(* Logix 5000 project; controller OWF Emulate 5570 rev 30.12; software revision 30.00; part 8 of 21 *)
(* tags used below, declared in another part *)
   OWF_Add_c : DINT;
   OWF_Input : DINT[16];
   OWF_Result : DINT[17];
(* MainProgram, continued *)

   	End_If;
   	If OWF_Input[7].[22] Then
   		OWF_Result[0]:=OWF_Result[0] + 480646434+OWF_Add_c;
   		OWF_Add_c.0:=OWF_Result[0].31;
   		OWF_Result[0].31:=0;
   		OWF_Result[1]:=OWF_Result[1] + 114796889+OWF_Add_c;
   		OWF_Add_c.1:=OWF_Result[1].31;
   		OWF_Result[1].31:=0;
   		OWF_Result[2]:=OWF_Result[2] + 808245238+OWF_Add_c;
   		OWF_Add_c.2:=OWF_Result[2].31;
   		OWF_Result[2].31:=0;
   		OWF_Result[3]:=OWF_Result[3] + 1045553390+OWF_Add_c;
   		OWF_Add_c.3:=OWF_Result[3].31;
   		OWF_Result[3].31:=0;
   		OWF_Result[4]:=OWF_Result[4] + 1347272097+OWF_Add_c;
   		OWF_Add_c.4:=OWF_Result[4].31;
   		OWF_Result[4].31:=0;
   		OWF_Result[5]:=OWF_Result[5] + 212393883+OWF_Add_c;
   		OWF_Add_c.5:=OWF_Result[5].31;
   		OWF_Result[5].31:=0;
   		OWF_Result[6]:=OWF_Result[6] + 833811458+OWF_Add_c;
   		OWF_Add_c.6:=OWF_Result[6].31;
   		OWF_Result[6].31:=0;
   		OWF_Result[7]:=OWF_Result[7] + 657498953+OWF_Add_c;
   		OWF_Add_c.7:=OWF_Result[7].31;
   		OWF_Result[7].31:=0;
   		OWF_Result[8]:=OWF_Result[8] + 1633172185+OWF_Add_c;
   		OWF_Add_c.8:=OWF_Result[8].31;
   		OWF_Result[8].31:=0;
   		OWF_Result[9]:=OWF_Result[9] + 109189510+OWF_Add_c;
   		OWF_Add_c.9:=OWF_Result[9].31;
   		OWF_Result[9].31:=0;
   		OWF_Result[10]:=OWF_Result[10] + 1987125799+OWF_Add_c;
   		OWF_Add_c.10:=OWF_Result[10].31;
   		OWF_Result[10].31:=0;
   		OWF_Result[11]:=OWF_Result[11] + 790477840+OWF_Add_c;
   		OWF_Add_c.11:=OWF_Result[11].31;
   		OWF_Result[11].31:=0;
   		OWF_Result[12]:=OWF_Result[12] + 1317536711+OWF_Add_c;
   		OWF_Add_c.12:=OWF_Result[12].31;
   		OWF_Result[12].31:=0;
   	End_If;
   	If OWF_Input[7].[23] Then
   		OWF_Result[0]:=OWF_Result[0] + 740299143+OWF_Add_c;
   		OWF_Add_c.0:=OWF_Result[0].31;
   		OWF_Result[0].31:=0;
   		OWF_Result[1]:=OWF_Result[1] + 289363045+OWF_Add_c;
   		OWF_Add_c.1:=OWF_Result[1].31;
   		OWF_Result[1].31:=0;
   		OWF_Result[2]:=OWF_Result[2] + 506118578+OWF_Add_c;
   		OWF_Add_c.2:=OWF_Result[2].31;
   		OWF_Result[2].31:=0;
   		OWF_Result[3]:=OWF_Result[3] + 1440714184+OWF_Add_c;
   		OWF_Add_c.3:=OWF_Result[3].31;
   		OWF_Result[3].31:=0;
   		OWF_Result[4]:=OWF_Result[4] + 1773567421+OWF_Add_c;
   		OWF_Add_c.4:=OWF_Result[4].31;
   		OWF_Result[4].31:=0;
   		OWF_Result[5]:=OWF_Result[5] + 1795348463+OWF_Add_c;
   		OWF_Add_c.5:=OWF_Result[5].31;
   		OWF_Result[5].31:=0;
   		OWF_Result[6]:=OWF_Result[6] + 1980498485+OWF_Add_c;
   		OWF_Add_c.6:=OWF_Result[6].31;
   		OWF_Result[6].31:=0;
   		OWF_Result[7]:=OWF_Result[7] + 308789052+OWF_Add_c;
   		OWF_Add_c.7:=OWF_Result[7].31;
   		OWF_Result[7].31:=0;
   		OWF_Result[8]:=OWF_Result[8] + 1048758798+OWF_Add_c;
   		OWF_Add_c.8:=OWF_Result[8].31;
   		OWF_Result[8].31:=0;
   		OWF_Result[9]:=OWF_Result[9] + 916377049+OWF_Add_c;
   		OWF_Add_c.9:=OWF_Result[9].31;
   		OWF_Result[9].31:=0;
   		OWF_Result[10]:=OWF_Result[10] + 502789876+OWF_Add_c;
   		OWF_Add_c.10:=OWF_Result[10].31;
   		OWF_Result[10].31:=0;
   		OWF_Result[11]:=OWF_Result[11] + 629743481+OWF_Add_c;
   		OWF_Add_c.11:=OWF_Result[11].31;
   		OWF_Result[11].31:=0;
   		OWF_Result[12]:=OWF_Result[12] + 1676079784+OWF_Add_c;
   		OWF_Add_c.12:=OWF_Result[12].31;
   		OWF_Result[12].31:=0;
   	End_If;
   	If OWF_Input[7].[24] Then
   		OWF_Result[0]:=OWF_Result[0] + 978983842+OWF_Add_c;
   		OWF_Add_c.0:=OWF_Result[0].31;
   		OWF_Result[0].31:=0;
   		OWF_Result[1]:=OWF_Result[1] + 184076912+OWF_Add_c;
   		OWF_Add_c.1:=OWF_Result[1].31;
   		OWF_Result[1].31:=0;
   		OWF_Result[2]:=OWF_Result[2] + 18075719+OWF_Add_c;
   		OWF_Add_c.2:=OWF_Result[2].31;
   		OWF_Result[2].31:=0;
   		OWF_Result[3]:=OWF_Result[3] + 1672505732+OWF_Add_c;
   		OWF_Add_c.3:=OWF_Result[3].31;
   		OWF_Result[3].31:=0;
   		OWF_Result[4]:=OWF_Result[4] + 1803238491+OWF_Add_c;
   		OWF_Add_c.4:=OWF_Result[4].31;
   		OWF_Result[4].31:=0;
   		OWF_Result[5]:=OWF_Result[5] + 1332716281+OWF_Add_c;
   		OWF_Add_c.5:=OWF_Result[5].31;
   		OWF_Result[5].31:=0;
   		OWF_Result[6]:=OWF_Result[6] + 633027607+OWF_Add_c;
   		OWF_Add_c.6:=OWF_Result[6].31;
   		OWF_Result[6].31:=0;
   		OWF_Result[7]:=OWF_Result[7] + 1542211604+OWF_Add_c;
   		OWF_Add_c.7:=OWF_Result[7].31;
   		OWF_Result[7].31:=0;
   		OWF_Result[8]:=OWF_Result[8] + 716891059+OWF_Add_c;
   		OWF_Add_c.8:=OWF_Result[8].31;
   		OWF_Result[8].31:=0;
   		OWF_Result[9]:=OWF_Result[9] + 1337341351+OWF_Add_c;
   		OWF_Add_c.9:=OWF_Result[9].31;
   		OWF_Result[9].31:=0;
   		OWF_Result[10]:=OWF_Result[10] + 1718317461+OWF_Add_c;
   		OWF_Add_c.10:=OWF_Result[10].31;
   		OWF_Result[10].31:=0;
   		OWF_Result[11]:=OWF_Result[11] + 759267344+OWF_Add_c;
   		OWF_Add_c.11:=OWF_Result[11].31;
   		OWF_Result[11].31:=0;
   		OWF_Result[12]:=OWF_Result[12] + 1222721366+OWF_Add_c;
   		OWF_Add_c.12:=OWF_Result[12].31;
   		OWF_Result[12].31:=0;
   	End_If;
   	If OWF_Input[7].[25] Then
   		OWF_Result[0]:=OWF_Result[0] + 1210573640+OWF_Add_c;
   		OWF_Add_c.0:=OWF_Result[0].31;
   		OWF_Result[0].31:=0;
   		OWF_Result[1]:=OWF_Result[1] + 1066502865+OWF_Add_c;
   		OWF_Add_c.1:=OWF_Result[1].31;
   		OWF_Result[1].31:=0;
   		OWF_Result[2]:=OWF_Result[2] + 20470411+OWF_Add_c;
   		OWF_Add_c.2:=OWF_Result[2].31;
   		OWF_Result[2].31:=0;
   		OWF_Result[3]:=OWF_Result[3] + 526137192+OWF_Add_c;
   		OWF_Add_c.3:=OWF_Result[3].31;
   		OWF_Result[3].31:=0;
   		OWF_Result[4]:=OWF_Result[4] + 428761318+OWF_Add_c;
   		OWF_Add_c.4:=OWF_Result[4].31;
   		OWF_Result[4].31:=0;
   		OWF_Result[5]:=OWF_Result[5] + 666284081+OWF_Add_c;
   		OWF_Add_c.5:=OWF_Result[5].31;
   		OWF_Result[5].31:=0;
   		OWF_Result[6]:=OWF_Result[6] + 787646009+OWF_Add_c;
   		OWF_Add_c.6:=OWF_Result[6].31;
   		OWF_Result[6].31:=0;
   		OWF_Result[7]:=OWF_Result[7] + 1465565705+OWF_Add_c;
   		OWF_Add_c.7:=OWF_Result[7].31;
   		OWF_Result[7].31:=0;
   		OWF_Result[8]:=OWF_Result[8] + 2117689109+OWF_Add_c;
   		OWF_Add_c.8:=OWF_Result[8].31;
   		OWF_Result[8].31:=0;
   		OWF_Result[9]:=OWF_Result[9] + 1455398601+OWF_Add_c;
   		OWF_Add_c.9:=OWF_Result[9].31;
   		OWF_Result[9].31:=0;
   		OWF_Result[10]:=OWF_Result[10] + 732503870+OWF_Add_c;
   		OWF_Add_c.10:=OWF_Result[10].31;
   		OWF_Result[10].31:=0;
   		OWF_Result[11]:=OWF_Result[11] + 1389721484+OWF_Add_c;
   		OWF_Add_c.11:=OWF_Result[11].31;
   		OWF_Result[11].31:=0;
   		OWF_Result[12]:=OWF_Result[12] + 1051435137+OWF_Add_c;
   		OWF_Add_c.12:=OWF_Result[12].31;
   		OWF_Result[12].31:=0;
   	End_If;
   	If OWF_Input[7].[26] Then
   		OWF_Result[0]:=OWF_Result[0] + 1093740877+OWF_Add_c;
   		OWF_Add_c.0:=OWF_Result[0].31;
   		OWF_Result[0].31:=0;
   		OWF_Result[1]:=OWF_Result[1] + 1926933030+OWF_Add_c;
   		OWF_Add_c.1:=OWF_Result[1].31;
   		OWF_Result[1].31:=0;
   		OWF_Result[2]:=OWF_Result[2] + 2048297708+OWF_Add_c;
   		OWF_Add_c.2:=OWF_Result[2].31;
   		OWF_Result[2].31:=0;
   		OWF_Result[3]:=OWF_Result[3] + 1774994164+OWF_Add_c;
   		OWF_Add_c.3:=OWF_Result[3].31;
   		OWF_Result[3].31:=0;
   		OWF_Result[4]:=OWF_Result[4] + 100463613+OWF_Add_c;
   		OWF_Add_c.4:=OWF_Result[4].31;
   		OWF_Result[4].31:=0;
   		OWF_Result[5]:=OWF_Result[5] + 1811813667+OWF_Add_c;
   		OWF_Add_c.5:=OWF_Result[5].31;
   		OWF_Result[5].31:=0;
   		OWF_Result[6]:=OWF_Result[6] + 1209213066+OWF_Add_c;
   		OWF_Add_c.6:=OWF_Result[6].31;
   		OWF_Result[6].31:=0;
   		OWF_Result[7]:=OWF_Result[7] + 1269950558+OWF_Add_c;
   		OWF_Add_c.7:=OWF_Result[7].31;
   		OWF_Result[7].31:=0;
   		OWF_Result[8]:=OWF_Result[8] + 624695169+OWF_Add_c;
   		OWF_Add_c.8:=OWF_Result[8].31;
   		OWF_Result[8].31:=0;
   		OWF_Result[9]:=OWF_Result[9] + 1916749071+OWF_Add_c;
   		OWF_Add_c.9:=OWF_Result[9].31;
   		OWF_Result[9].31:=0;
   		OWF_Result[10]:=OWF_Result[10] + 1775084911+OWF_Add_c;
   		OWF_Add_c.10:=OWF_Result[10].31;
   		OWF_Result[10].31:=0;
   		OWF_Result[11]:=OWF_Result[11] + 1305211684+OWF_Add_c;
   		OWF_Add_c.11:=OWF_Result[11].31;
   		OWF_Result[11].31:=0;
   		OWF_Result[12]:=OWF_Result[12] + 546822773+OWF_Add_c;
   		OWF_Add_c.12:=OWF_Result[12].31;
   		OWF_Result[12].31:=0;
   	End_If;
   	If OWF_Input[7].[27] Then
   		OWF_Result[0]:=OWF_Result[0] + 859091503+OWF_Add_c;
   		OWF_Add_c.0:=OWF_Result[0].31;
   		OWF_Result[0].31:=0;
   		OWF_Result[1]:=OWF_Result[1] + 734881955+OWF_Add_c;
   		OWF_Add_c.1:=OWF_Result[1].31;
   		OWF_Result[1].31:=0;
   		OWF_Result[2]:=OWF_Result[2] + 2112245734+OWF_Add_c;
   		OWF_Add_c.2:=OWF_Result[2].31;
   		OWF_Result[2].31:=0;
   		OWF_Result[3]:=OWF_Result[3] + 821086543+OWF_Add_c;
   		OWF_Add_c.3:=OWF_Result[3].31;
   		OWF_Result[3].31:=0;
   		OWF_Result[4]:=OWF_Result[4] + 172634749+OWF_Add_c;
   		OWF_Add_c.4:=OWF_Result[4].31;
   		OWF_Result[4].31:=0;
   		OWF_Result[5]:=OWF_Result[5] + 1640326127+OWF_Add_c;
   		OWF_Add_c.5:=OWF_Result[5].31;
   		OWF_Result[5].31:=0;
   		OWF_Result[6]:=OWF_Result[6] + 90813347+OWF_Add_c;
   		OWF_Add_c.6:=OWF_Result[6].31;
   		OWF_Result[6].31:=0;
   		OWF_Result[7]:=OWF_Result[7] + 375324933+OWF_Add_c;
   		OWF_Add_c.7:=OWF_Result[7].31;
   		OWF_Result[7].31:=0;
   		OWF_Result[8]:=OWF_Result[8] + 734165162+OWF_Add_c;
   		OWF_Add_c.8:=OWF_Result[8].31;
   		OWF_Result[8].31:=0;
   		OWF_Result[9]:=OWF_Result[9] + 1211646497+OWF_Add_c;
   		OWF_Add_c.9:=OWF_Result[9].31;
   		OWF_Result[9].31:=0;
   		OWF_Result[10]:=OWF_Result[10] + 243057850+OWF_Add_c;
   		OWF_Add_c.10:=OWF_Result[10].31;
   		OWF_Result[10].31:=0;
   		OWF_Result[11]:=OWF_Result[11] + 2097424801+OWF_Add_c;
   		OWF_Add_c.11:=OWF_Result[11].31;
   		OWF_Result[11].31:=0;
   		OWF_Result[12]:=OWF_Result[12] + 609462236+OWF_Add_c;
   		OWF_Add_c.12:=OWF_Result[12].31;
   		OWF_Result[12].31:=0;
   	End_If;
   	If OWF_Input[7].[28] Then
   		OWF_Result[0]:=OWF_Result[0] + 1748630085+OWF_Add_c;
   		OWF_Add_c.0:=OWF_Result[0].31;
   		OWF_Result[0].31:=0;
   		OWF_Result[1]:=OWF_Result[1] + 218806354+OWF_Add_c;
   		OWF_Add_c.1:=OWF_Result[1].31;
   		OWF_Result[1].31:=0;
   		OWF_Result[2]:=OWF_Result[2] + 596066578+OWF_Add_c;
   		OWF_Add_c.2:=OWF_Result[2].31;
   		OWF_Result[2].31:=0;
   		OWF_Result[3]:=OWF_Result[3] + 1279944685+OWF_Add_c;
   		OWF_Add_c.3:=OWF_Result[3].31;
   		OWF_Result[3].31:=0;
   		OWF_Result[4]:=OWF_Result[4] + 798939716+OWF_Add_c;
   		OWF_Add_c.4:=OWF_Result[4].31;
   		OWF_Result[4].31:=0;
   		OWF_Result[5]:=OWF_Result[5] + 1193007422+OWF_Add_c;
   		OWF_Add_c.5:=OWF_Result[5].31;
   		OWF_Result[5].31:=0;
   		OWF_Result[6]:=OWF_Result[6] + 718950431+OWF_Add_c;
   		OWF_Add_c.6:=OWF_Result[6].31;
   		OWF_Result[6].31:=0;
   		OWF_Result[7]:=OWF_Result[7] + 576120375+OWF_Add_c;
   		OWF_Add_c.7:=OWF_Result[7].31;
   		OWF_Result[7].31:=0;
   		OWF_Result[8]:=OWF_Result[8] + 1793230797+OWF_Add_c;
   		OWF_Add_c.8:=OWF_Result[8].31;
   		OWF_Result[8].31:=0;
   		OWF_Result[9]:=OWF_Result[9] + 482018913+OWF_Add_c;
   		OWF_Add_c.9:=OWF_Result[9].31;
   		OWF_Result[9].31:=0;
   		OWF_Result[10]:=OWF_Result[10] + 434876156+OWF_Add_c;
   		OWF_Add_c.10:=OWF_Result[10].31;
   		OWF_Result[10].31:=0;
   		OWF_Result[11]:=OWF_Result[11] + 228585162+OWF_Add_c;
   		OWF_Add_c.11:=OWF_Result[11].31;
   		OWF_Result[11].31:=0;
   		OWF_Result[12]:=OWF_Result[12] + 868694246+OWF_Add_c;
   		OWF_Add_c.12:=OWF_Result[12].31;
   		OWF_Result[12].31:=0;
   	End_If;
   	If OWF_Input[7].[29] Then
   		OWF_Result[0]:=OWF_Result[0] + 1193337411+OWF_Add_c;
   		OWF_Add_c.0:=OWF_Result[0].31;
   		OWF_Result[0].31:=0;
   		OWF_Result[1]:=OWF_Result[1] + 1791500938+OWF_Add_c;
   		OWF_Add_c.1:=OWF_Result[1].31;
   		OWF_Result[1].31:=0;
   		OWF_Result[2]:=OWF_Result[2] + 518096871+OWF_Add_c;
   		OWF_Add_c.2:=OWF_Result[2].31;
   		OWF_Result[2].31:=0;
   		OWF_Result[3]:=OWF_Result[3] + 1495747504+OWF_Add_c;
   		OWF_Add_c.3:=OWF_Result[3].31;
   		OWF_Result[3].31:=0;
   		OWF_Result[4]:=OWF_Result[4] + 1777942201+OWF_Add_c;
   		OWF_Add_c.4:=OWF_Result[4].31;
   		OWF_Result[4].31:=0;
   		OWF_Result[5]:=OWF_Result[5] + 275225992+OWF_Add_c;
   		OWF_Add_c.5:=OWF_Result[5].31;
   		OWF_Result[5].31:=0;
   		OWF_Result[6]:=OWF_Result[6] + 826164955+OWF_Add_c;
   		OWF_Add_c.6:=OWF_Result[6].31;
   		OWF_Result[6].31:=0;
   		OWF_Result[7]:=OWF_Result[7] + 157561222+OWF_Add_c;
   		OWF_Add_c.7:=OWF_Result[7].31;
   		OWF_Result[7].31:=0;
   		OWF_Result[8]:=OWF_Result[8] + 1558104080+OWF_Add_c;
   		OWF_Add_c.8:=OWF_Result[8].31;
   		OWF_Result[8].31:=0;
   		OWF_Result[9]:=OWF_Result[9] + 1972530605+OWF_Add_c;
   		OWF_Add_c.9:=OWF_Result[9].31;
   		OWF_Result[9].31:=0;
   		OWF_Result[10]:=OWF_Result[10] + 61824397+OWF_Add_c;
   		OWF_Add_c.10:=OWF_Result[10].31;
   		OWF_Result[10].31:=0;
   		OWF_Result[11]:=OWF_Result[11] + 1231944572+OWF_Add_c;
   		OWF_Add_c.11:=OWF_Result[11].31;
   		OWF_Result[11].31:=0;
   		OWF_Result[12]:=OWF_Result[12] + 1095576086+OWF_Add_c;
   		OWF_Add_c.12:=OWF_Result[12].31;
   		OWF_Result[12].31:=0;
   	End_If;
   	If OWF_Input[7].[30] Then
   		OWF_Result[0]:=OWF_Result[0] + 235927346+OWF_Add_c;
   		OWF_Add_c.0:=OWF_Result[0].31;
   		OWF_Result[0].31:=0;
   		OWF_Result[1]:=OWF_Result[1] + 405435054+OWF_Add_c;
   		OWF_Add_c.1:=OWF_Result[1].31;
   		OWF_Result[1].31:=0;
   		OWF_Result[2]:=OWF_Result[2] + 310760218+OWF_Add_c;
   		OWF_Add_c.2:=OWF_Result[2].31;
   		OWF_Result[2].31:=0;
   		OWF_Result[3]:=OWF_Result[3] + 1004598596+OWF_Add_c;
   		OWF_Add_c.3:=OWF_Result[3].31;
   		OWF_Result[3].31:=0;
   		OWF_Result[4]:=OWF_Result[4] + 636478930+OWF_Add_c;
   		OWF_Add_c.4:=OWF_Result[4].31;
   		OWF_Result[4].31:=0;
   		OWF_Result[5]:=OWF_Result[5] + 1964479220+OWF_Add_c;
   		OWF_Add_c.5:=OWF_Result[5].31;
   		OWF_Result[5].31:=0;
   		OWF_Result[6]:=OWF_Result[6] + 391120426+OWF_Add_c;
   		OWF_Add_c.6:=OWF_Result[6].31;
   		OWF_Result[6].31:=0;
   		OWF_Result[7]:=OWF_Result[7] + 953930079+OWF_Add_c;
   		OWF_Add_c.7:=OWF_Result[7].31;
   		OWF_Result[7].31:=0;
   		OWF_Result[8]:=OWF_Result[8] + 1444849706+OWF_Add_c;
   		OWF_Add_c.8:=OWF_Result[8].31;
   		OWF_Result[8].31:=0;
   		OWF_Result[9]:=OWF_Result[9] + 1419197967+OWF_Add_c;
   		OWF_Add_c.9:=OWF_Result[9].31;
   		OWF_Result[9].31:=0;
   		OWF_Result[10]:=OWF_Result[10] + 84707091+OWF_Add_c;
   		OWF_Add_c.10:=OWF_Result[10].31;
   		OWF_Result[10].31:=0;
   		OWF_Result[11]:=OWF_Result[11] + 727669007+OWF_Add_c;
   		OWF_Add_c.11:=OWF_Result[11].31;
   		OWF_Result[11].31:=0;
   		OWF_Result[12]:=OWF_Result[12] + 242116771+OWF_Add_c;
   		OWF_Add_c.12:=OWF_Result[12].31;
   		OWF_Result[12].31:=0;
   	End_If;
   	If OWF_Input[7].[31] Then
   		OWF_Result[0]:=OWF_Result[0] + 415305185+OWF_Add_c;
   		OWF_Add_c.0:=OWF_Result[0].31;
   		OWF_Result[0].31:=0;
   		OWF_Result[1]:=OWF_Result[1] + 1993683176+OWF_Add_c;
   		OWF_Add_c.1:=OWF_Result[1].31;
   		OWF_Result[1].31:=0;
   		OWF_Result[2]:=OWF_Result[2] + 2081036556+OWF_Add_c;
   		OWF_Add_c.2:=OWF_Result[2].31;
   		OWF_Result[2].31:=0;
   		OWF_Result[3]:=OWF_Result[3] + 926823350+OWF_Add_c;
   		OWF_Add_c.3:=OWF_Result[3].31;
   		OWF_Result[3].31:=0;
   		OWF_Result[4]:=OWF_Result[4] + 426179276+OWF_Add_c;
   		OWF_Add_c.4:=OWF_Result[4].31;
   		OWF_Result[4].31:=0;
   		OWF_Result[5]:=OWF_Result[5] + 2096822006+OWF_Add_c;
   		OWF_Add_c.5:=OWF_Result[5].31;
   		OWF_Result[5].31:=0;
   		OWF_Result[6]:=OWF_Result[6] + 1622929595+OWF_Add_c;
   		OWF_Add_c.6:=OWF_Result[6].31;
   		OWF_Result[6].31:=0;
   		OWF_Result[7]:=OWF_Result[7] + 1783463523+OWF_Add_c;
   		OWF_Add_c.7:=OWF_Result[7].31;
   		OWF_Result[7].31:=0;
   		OWF_Result[8]:=OWF_Result[8] + 1221615485+OWF_Add_c;
   		OWF_Add_c.8:=OWF_Result[8].31;
   		OWF_Result[8].31:=0;
   		OWF_Result[9]:=OWF_Result[9] + 783241525+OWF_Add_c;
   		OWF_Add_c.9:=OWF_Result[9].31;
   		OWF_Result[9].31:=0;
   		OWF_Result[10]:=OWF_Result[10] + 13423679+OWF_Add_c;
   		OWF_Add_c.10:=OWF_Result[10].31;
   		OWF_Result[10].31:=0;
   		OWF_Result[11]:=OWF_Result[11] + 552970833+OWF_Add_c;
   		OWF_Add_c.11:=OWF_Result[11].31;
   		OWF_Result[11].31:=0;
   		OWF_Result[12]:=OWF_Result[12] + 1709245061+OWF_Add_c;
   		OWF_Add_c.12:=OWF_Result[12].31;
   		OWF_Result[12].31:=0;
   	End_If;
   	If OWF_Input[8].[0] Then
   		OWF_Result[0]:=OWF_Result[0] + 1733835665+OWF_Add_c;
   		OWF_Add_c.0:=OWF_Result[0].31;
   		OWF_Result[0].31:=0;
   		OWF_Result[1]:=OWF_Result[1] + 916519587+OWF_Add_c;
   		OWF_Add_c.1:=OWF_Result[1].31;
   		OWF_Result[1].31:=0;
   		OWF_Result[2]:=OWF_Result[2] + 2058734345+OWF_Add_c;
   		OWF_Add_c.2:=OWF_Result[2].31;
   		OWF_Result[2].31:=0;
   		OWF_Result[3]:=OWF_Result[3] + 1314200972+OWF_Add_c;
   		OWF_Add_c.3:=OWF_Result[3].31;
   		OWF_Result[3].31:=0;
   		OWF_Result[4]:=OWF_Result[4] + 876718991+OWF_Add_c;
   		OWF_Add_c.4:=OWF_Result[4].31;
   		OWF_Result[4].31:=0;
   		OWF_Result[5]:=OWF_Result[5] + 5729275+OWF_Add_c;
   		OWF_Add_c.5:=OWF_Result[5].31;
   		OWF_Result[5].31:=0;
   		OWF_Result[6]:=OWF_Result[6] + 506795812+OWF_Add_c;
   		OWF_Add_c.6:=OWF_Result[6].31;
   		OWF_Result[6].31:=0;
   		OWF_Result[7]:=OWF_Result[7] + 722793935+OWF_Add_c;
   		OWF_Add_c.7:=OWF_Result[7].31;
   		OWF_Result[7].31:=0;
   		OWF_Result[8]:=OWF_Result[8] + 1119541514+OWF_Add_c;
   		OWF_Add_c.8:=OWF_Result[8].31;
   		OWF_Result[8].31:=0;
   		OWF_Result[9]:=OWF_Result[9] + 1442255024+OWF_Add_c;
   		OWF_Add_c.9:=OWF_Result[9].31;
   		OWF_Result[9].31:=0;
   		OWF_Result[10]:=OWF_Result[10] + 10828735+OWF_Add_c;
   		OWF_Add_c.10:=OWF_Result[10].31;
   		OWF_Result[10].31:=0;
   		OWF_Result[11]:=OWF_Result[11] + 1845527341+OWF_Add_c;
   		OWF_Add_c.11:=OWF_Result[11].31;
   		OWF_Result[11].31:=0;
   		OWF_Result[12]:=OWF_Result[12] + 864596063+OWF_Add_c;
   		OWF_Add_c.12:=OWF_Result[12].31;
   		OWF_Result[12].31:=0;
   	End_If;
   	If OWF_Input[8].[1] Then
   		OWF_Result[0]:=OWF_Result[0] + 176336629+OWF_Add_c;
   		OWF_Add_c.0:=OWF_Result[0].31;
   		OWF_Result[0].31:=0;
   		OWF_Result[1]:=OWF_Result[1] + 46344304+OWF_Add_c;
   		OWF_Add_c.1:=OWF_Result[1].31;
   		OWF_Result[1].31:=0;
   		OWF_Result[2]:=OWF_Result[2] + 58822969+OWF_Add_c;
   		OWF_Add_c.2:=OWF_Result[2].31;
   		OWF_Result[2].31:=0;
   		OWF_Result[3]:=OWF_Result[3] + 1869389297+OWF_Add_c;
   		OWF_Add_c.3:=OWF_Result[3].31;
   		OWF_Result[3].31:=0;
   		OWF_Result[4]:=OWF_Result[4] + 758725144+OWF_Add_c;
   		OWF_Add_c.4:=OWF_Result[4].31;
   		OWF_Result[4].31:=0;
   		OWF_Result[5]:=OWF_Result[5] + 1234591682+OWF_Add_c;
   		OWF_Add_c.5:=OWF_Result[5].31;
   		OWF_Result[5].31:=0;
   		OWF_Result[6]:=OWF_Result[6] + 2101460213+OWF_Add_c;
   		OWF_Add_c.6:=OWF_Result[6].31;
   		OWF_Result[6].31:=0;
   		OWF_Result[7]:=OWF_Result[7] + 189121499+OWF_Add_c;
   		OWF_Add_c.7:=OWF_Result[7].31;
   		OWF_Result[7].31:=0;
   		OWF_Result[8]:=OWF_Result[8] + 1567832861+OWF_Add_c;
   		OWF_Add_c.8:=OWF_Result[8].31;
   		OWF_Result[8].31:=0;
   		OWF_Result[9]:=OWF_Result[9] + 50878325+OWF_Add_c;
   		OWF_Add_c.9:=OWF_Result[9].31;
   		OWF_Result[9].31:=0;
   		OWF_Result[10]:=OWF_Result[10] + 380406108+OWF_Add_c;
   		OWF_Add_c.10:=OWF_Result[10].31;
   		OWF_Result[10].31:=0;
   		OWF_Result[11]:=OWF_Result[11] + 119007880+OWF_Add_c;
   		OWF_Add_c.11:=OWF_Result[11].31;
   		OWF_Result[11].31:=0;
   		OWF_Result[12]:=OWF_Result[12] + 1980093434+OWF_Add_c;
   		OWF_Add_c.12:=OWF_Result[12].31;
   		OWF_Result[12].31:=0;
   	End_If;
   	If OWF_Input[8].[2] Then
   		OWF_Result[0]:=OWF_Result[0] + 928675896+OWF_Add_c;
   		OWF_Add_c.0:=OWF_Result[0].31;
   		OWF_Result[0].31:=0;
   		OWF_Result[1]:=OWF_Result[1] + 505177878+OWF_Add_c;
   		OWF_Add_c.1:=OWF_Result[1].31;
   		OWF_Result[1].31:=0;
   		OWF_Result[2]:=OWF_Result[2] + 1750158252+OWF_Add_c;
   		OWF_Add_c.2:=OWF_Result[2].31;
   		OWF_Result[2].31:=0;
   		OWF_Result[3]:=OWF_Result[3] + 509803710+OWF_Add_c;
   		OWF_Add_c.3:=OWF_Result[3].31;
   		OWF_Result[3].31:=0;
   		OWF_Result[4]:=OWF_Result[4] + 517535777+OWF_Add_c;
   		OWF_Add_c.4:=OWF_Result[4].31;
   		OWF_Result[4].31:=0;
   		OWF_Result[5]:=OWF_Result[5] + 1876669972+OWF_Add_c;
   		OWF_Add_c.5:=OWF_Result[5].31;
   		OWF_Result[5].31:=0;
   		OWF_Result[6]:=OWF_Result[6] + 1296281635+OWF_Add_c;
   		OWF_Add_c.6:=OWF_Result[6].31;
   		OWF_Result[6].31:=0;
   		OWF_Result[7]:=OWF_Result[7] + 196070166+OWF_Add_c;
   		OWF_Add_c.7:=OWF_Result[7].31;
   		OWF_Result[7].31:=0;
   		OWF_Result[8]:=OWF_Result[8] + 1491248578+OWF_Add_c;
   		OWF_Add_c.8:=OWF_Result[8].31;
   		OWF_Result[8].31:=0;
   		OWF_Result[9]:=OWF_Result[9] + 308195660+OWF_Add_c;
   		OWF_Add_c.9:=OWF_Result[9].31;
   		OWF_Result[9].31:=0;
   		OWF_Result[10]:=OWF_Result[10] + 493476372+OWF_Add_c;
   		OWF_Add_c.10:=OWF_Result[10].31;
   		OWF_Result[10].31:=0;
   		OWF_Result[11]:=OWF_Result[11] + 1546260645+OWF_Add_c;
   		OWF_Add_c.11:=OWF_Result[11].31;
   		OWF_Result[11].31:=0;
   		OWF_Result[12]:=OWF_Result[12] + 1306588125+OWF_Add_c;
   		OWF_Add_c.12:=OWF_Result[12].31;
   		OWF_Result[12].31:=0;
   	End_If;
   	If OWF_Input[8].[3] Then
   		OWF_Result[0]:=OWF_Result[0] + 181953250+OWF_Add_c;
   		OWF_Add_c.0:=OWF_Result[0].31;
   		OWF_Result[0].31:=0;
   		OWF_Result[1]:=OWF_Result[1] + 790129216+OWF_Add_c;
   		OWF_Add_c.1:=OWF_Result[1].31;
   		OWF_Result[1].31:=0;
   		OWF_Result[2]:=OWF_Result[2] + 52204497+OWF_Add_c;
   		OWF_Add_c.2:=OWF_Result[2].31;
   		OWF_Result[2].31:=0;
   		OWF_Result[3]:=OWF_Result[3] + 1999525053+OWF_Add_c;
   		OWF_Add_c.3:=OWF_Result[3].31;
   		OWF_Result[3].31:=0;
   		OWF_Result[4]:=OWF_Result[4] + 439204566+OWF_Add_c;
   		OWF_Add_c.4:=OWF_Result[4].31;
   		OWF_Result[4].31:=0;
   		OWF_Result[5]:=OWF_Result[5] + 770505550+OWF_Add_c;
   		OWF_Add_c.5:=OWF_Result[5].31;
   		OWF_Result[5].31:=0;
   		OWF_Result[6]:=OWF_Result[6] + 1508348621+OWF_Add_c;
   		OWF_Add_c.6:=OWF_Result[6].31;
   		OWF_Result[6].31:=0;
   		OWF_Result[7]:=OWF_Result[7] + 150288603+OWF_Add_c;
   		OWF_Add_c.7:=OWF_Result[7].31;
   		OWF_Result[7].31:=0;
   		OWF_Result[8]:=OWF_Result[8] + 908594+OWF_Add_c;
   		OWF_Add_c.8:=OWF_Result[8].31;
   		OWF_Result[8].31:=0;
   		OWF_Result[9]:=OWF_Result[9] + 938186794+OWF_Add_c;
   		OWF_Add_c.9:=OWF_Result[9].31;
   		OWF_Result[9].31:=0;
   		OWF_Result[10]:=OWF_Result[10] + 1270944269+OWF_Add_c;
   		OWF_Add_c.10:=OWF_Result[10].31;
   		OWF_Result[10].31:=0;
   		OWF_Result[11]:=OWF_Result[11] + 707941313+OWF_Add_c;
   		OWF_Add_c.11:=OWF_Result[11].31;
   		OWF_Result[11].31:=0;
   		OWF_Result[12]:=OWF_Result[12] + 182040987+OWF_Add_c;
   		OWF_Add_c.12:=OWF_Result[12].31;
   		OWF_Result[12].31:=0;
   	End_If;
   	If OWF_Input[8].[4] Then
   		OWF_Result[0]:=OWF_Result[0] + 35324931+OWF_Add_c;
   		OWF_Add_c.0:=OWF_Result[0].31;
   		OWF_Result[0].31:=0;
   		OWF_Result[1]:=OWF_Result[1] + 390808332+OWF_Add_c;
   		OWF_Add_c.1:=OWF_Result[1].31;
   		OWF_Result[1].31:=0;
   		OWF_Result[2]:=OWF_Result[2] + 831042246+OWF_Add_c;
   		OWF_Add_c.2:=OWF_Result[2].31;
   		OWF_Result[2].31:=0;
   		OWF_Result[3]:=OWF_Result[3] + 1714707837+OWF_Add_c;
   		OWF_Add_c.3:=OWF_Result[3].31;
   		OWF_Result[3].31:=0;
   		OWF_Result[4]:=OWF_Result[4] + 895947097+OWF_Add_c;
   		OWF_Add_c.4:=OWF_Result[4].31;
   		OWF_Result[4].31:=0;
   		OWF_Result[5]:=OWF_Result[5] + 324590523+OWF_Add_c;
   		OWF_Add_c.5:=OWF_Result[5].31;
   		OWF_Result[5].31:=0;
   		OWF_Result[6]:=OWF_Result[6] + 1399448768+OWF_Add_c;
   		OWF_Add_c.6:=OWF_Result[6].31;
   		OWF_Result[6].31:=0;
   		OWF_Result[7]:=OWF_Result[7] + 1771562066+OWF_Add_c;
   		OWF_Add_c.7:=OWF_Result[7].31;
   		OWF_Result[7].31:=0;
   		OWF_Result[8]:=OWF_Result[8] + 2009853435+OWF_Add_c;
   		OWF_Add_c.8:=OWF_Result[8].31;
   		OWF_Result[8].31:=0;
   		OWF_Result[9]:=OWF_Result[9] + 1737076810+OWF_Add_c;
   		OWF_Add_c.9:=OWF_Result[9].31;
   		OWF_Result[9].31:=0;
   		OWF_Result[10]:=OWF_Result[10] + 327974283+OWF_Add_c;
   		OWF_Add_c.10:=OWF_Result[10].31;
   		OWF_Result[10].31:=0;
   		OWF_Result[11]:=OWF_Result[11] + 1336577511+OWF_Add_c;
   		OWF_Add_c.11:=OWF_Result[11].31;
   		OWF_Result[11].31:=0;
   		OWF_Result[12]:=OWF_Result[12] + 503968909+OWF_Add_c;
   		OWF_Add_c.12:=OWF_Result[12].31;
   		OWF_Result[12].31:=0;
   	End_If;
   	If OWF_Input[8].[5] Then
   		OWF_Result[0]:=OWF_Result[0] + 1606715828+OWF_Add_c;
   		OWF_Add_c.0:=OWF_Result[0].31;
   		OWF_Result[0].31:=0;
   		OWF_Result[1]:=OWF_Result[1] + 60669240+OWF_Add_c;
   		OWF_Add_c.1:=OWF_Result[1].31;
   		OWF_Result[1].31:=0;
   		OWF_Result[2]:=OWF_Result[2] + 2036856136+OWF_Add_c;
   		OWF_Add_c.2:=OWF_Result[2].31;
   		OWF_Result[2].31:=0;
   		OWF_Result[3]:=OWF_Result[3] + 853418547+OWF_Add_c;
   		OWF_Add_c.3:=OWF_Result[3].31;
   		OWF_Result[3].31:=0;
   		OWF_Result[4]:=OWF_Result[4] + 788881870+OWF_Add_c;
   		OWF_Add_c.4:=OWF_Result[4].31;
   		OWF_Result[4].31:=0;
   		OWF_Result[5]:=OWF_Result[5] + 1312511236+OWF_Add_c;
   		OWF_Add_c.5:=OWF_Result[5].31;
   		OWF_Result[5].31:=0;
   		OWF_Result[6]:=OWF_Result[6] + 825357085+OWF_Add_c;
   		OWF_Add_c.6:=OWF_Result[6].31;
   		OWF_Result[6].31:=0;
   		OWF_Result[7]:=OWF_Result[7] + 1908480029+OWF_Add_c;
   		OWF_Add_c.7:=OWF_Result[7].31;
   		OWF_Result[7].31:=0;
   		OWF_Result[8]:=OWF_Result[8] + 2103253624+OWF_Add_c;
   		OWF_Add_c.8:=OWF_Result[8].31;
   		OWF_Result[8].31:=0;
   		OWF_Result[9]:=OWF_Result[9] + 1523871832+OWF_Add_c;
   		OWF_Add_c.9:=OWF_Result[9].31;
   		OWF_Result[9].31:=0;
   		OWF_Result[10]:=OWF_Result[10] + 784833363+OWF_Add_c;
   		OWF_Add_c.10:=OWF_Result[10].31;
   		OWF_Result[10].31:=0;
   		OWF_Result[11]:=OWF_Result[11] + 1815265117+OWF_Add_c;
   		OWF_Add_c.11:=OWF_Result[11].31;
   		OWF_Result[11].31:=0;
   		OWF_Result[12]:=OWF_Result[12] + 1171080340+OWF_Add_c;
   		OWF_Add_c.12:=OWF_Result[12].31;
   		OWF_Result[12].31:=0;
   	End_If;
   	If OWF_Input[8].[6] Then
   		OWF_Result[0]:=OWF_Result[0] + 1062532440+OWF_Add_c;
   		OWF_Add_c.0:=OWF_Result[0].31;
   		OWF_Result[0].31:=0;
   		OWF_Result[1]:=OWF_Result[1] + 1730530273+OWF_Add_c;
   		OWF_Add_c.1:=OWF_Result[1].31;
   		OWF_Result[1].31:=0;
   		OWF_Result[2]:=OWF_Result[2] + 147317301+OWF_Add_c;
   		OWF_Add_c.2:=OWF_Result[2].31;
   		OWF_Result[2].31:=0;
   		OWF_Result[3]:=OWF_Result[3] + 1364210765+OWF_Add_c;
   		OWF_Add_c.3:=OWF_Result[3].31;
   		OWF_Result[3].31:=0;
   		OWF_Result[4]:=OWF_Result[4] + 952088146+OWF_Add_c;
   		OWF_Add_c.4:=OWF_Result[4].31;
   		OWF_Result[4].31:=0;
   		OWF_Result[5]:=OWF_Result[5] + 1315721657+OWF_Add_c;
   		OWF_Add_c.5:=OWF_Result[5].31;
   		OWF_Result[5].31:=0;
   		OWF_Result[6]:=OWF_Result[6] + 1051306675+OWF_Add_c;
   		OWF_Add_c.6:=OWF_Result[6].31;
   		OWF_Result[6].31:=0;
   		OWF_Result[7]:=OWF_Result[7] + 448836047+OWF_Add_c;
   		OWF_Add_c.7:=OWF_Result[7].31;
   		OWF_Result[7].31:=0;
   		OWF_Result[8]:=OWF_Result[8] + 89403910+OWF_Add_c;
   		OWF_Add_c.8:=OWF_Result[8].31;
   		OWF_Result[8].31:=0;
   		OWF_Result[9]:=OWF_Result[9] + 1093634171+OWF_Add_c;
   		OWF_Add_c.9:=OWF_Result[9].31;
   		OWF_Result[9].31:=0;
   		OWF_Result[10]:=OWF_Result[10] + 449471534+OWF_Add_c;
   		OWF_Add_c.10:=OWF_Result[10].31;
   		OWF_Result[10].31:=0;
   		OWF_Result[11]:=OWF_Result[11] + 60589753+OWF_Add_c;
   		OWF_Add_c.11:=OWF_Result[11].31;
   		OWF_Result[11].31:=0;
   		OWF_Result[12]:=OWF_Result[12] + 85142838+OWF_Add_c;
   		OWF_Add_c.12:=OWF_Result[12].31;
   		OWF_Result[12].31:=0;
   	End_If;
   	If OWF_Input[8].[7] Then
   		OWF_Result[0]:=OWF_Result[0] + 1687821066+OWF_Add_c;
   		OWF_Add_c.0:=OWF_Result[0].31;
   		OWF_Result[0].31:=0;
   		OWF_Result[1]:=OWF_Result[1] + 951544335+OWF_Add_c;
   		OWF_Add_c.1:=OWF_Result[1].31;
   		OWF_Result[1].31:=0;
   		OWF_Result[2]:=OWF_Result[2] + 1805920537+OWF_Add_c;
   		OWF_Add_c.2:=OWF_Result[2].31;
   		OWF_Result[2].31:=0;
   		OWF_Result[3]:=OWF_Result[3] + 714932068+OWF_Add_c;
   		OWF_Add_c.3:=OWF_Result[3].31;
   		OWF_Result[3].31:=0;
   		OWF_Result[4]:=OWF_Result[4] + 960609119+OWF_Add_c;
   		OWF_Add_c.4:=OWF_Result[4].31;
   		OWF_Result[4].31:=0;
   		OWF_Result[5]:=OWF_Result[5] + 1739410571+OWF_Add_c;
   		OWF_Add_c.5:=OWF_Result[5].31;
   		OWF_Result[5].31:=0;
   		OWF_Result[6]:=OWF_Result[6] + 1961837903+OWF_Add_c;
   		OWF_Add_c.6:=OWF_Result[6].31;
   		OWF_Result[6].31:=0;
   		OWF_Result[7]:=OWF_Result[7] + 901175212+OWF_Add_c;
   		OWF_Add_c.7:=OWF_Result[7].31;
   		OWF_Result[7].31:=0;
   		OWF_Result[8]:=OWF_Result[8] + 1803719590+OWF_Add_c;
   		OWF_Add_c.8:=OWF_Result[8].31;
   		OWF_Result[8].31:=0;
   		OWF_Result[9]:=OWF_Result[9] + 380747488+OWF_Add_c;
   		OWF_Add_c.9:=OWF_Result[9].31;
   		OWF_Result[9].31:=0;
   		OWF_Result[10]:=OWF_Result[10] + 2021367515+OWF_Add_c;
   		OWF_Add_c.10:=OWF_Result[10].31;
   		OWF_Result[10].31:=0;
   		OWF_Result[11]:=OWF_Result[11] + 1465559353+OWF_Add_c;
   		OWF_Add_c.11:=OWF_Result[11].31;
   		OWF_Result[11].31:=0;
   		OWF_Result[12]:=OWF_Result[12] + 1048087069+OWF_Add_c;
   		OWF_Add_c.12:=OWF_Result[12].31;
   		OWF_Result[12].31:=0;
   	End_If;
   	If OWF_Input[8].[8] Then
   		OWF_Result[0]:=OWF_Result[0] + 2094814625+OWF_Add_c;
   		OWF_Add_c.0:=OWF_Result[0].31;
   		OWF_Result[0].31:=0;
   		OWF_Result[1]:=OWF_Result[1] + 201453386+OWF_Add_c;
   		OWF_Add_c.1:=OWF_Result[1].31;
   		OWF_Result[1].31:=0;
   		OWF_Result[2]:=OWF_Result[2] + 1480082638+OWF_Add_c;
   		OWF_Add_c.2:=OWF_Result[2].31;
   		OWF_Result[2].31:=0;
   		OWF_Result[3]:=OWF_Result[3] + 1862215500+OWF_Add_c;
   		OWF_Add_c.3:=OWF_Result[3].31;
   		OWF_Result[3].31:=0;
   		OWF_Result[4]:=OWF_Result[4] + 1964016082+OWF_Add_c;
   		OWF_Add_c.4:=OWF_Result[4].31;
   		OWF_Result[4].31:=0;
   		OWF_Result[5]:=OWF_Result[5] + 1326978276+OWF_Add_c;
   		OWF_Add_c.5:=OWF_Result[5].31;
   		OWF_Result[5].31:=0;
   		OWF_Result[6]:=OWF_Result[6] + 453175292+OWF_Add_c;
   		OWF_Add_c.6:=OWF_Result[6].31;
   		OWF_Result[6].31:=0;
   		OWF_Result[7]:=OWF_Result[7] + 2101594815+OWF_Add_c;
   		OWF_Add_c.7:=OWF_Result[7].31;
   		OWF_Result[7].31:=0;
   		OWF_Result[8]:=OWF_Result[8] + 107115492+OWF_Add_c;
   		OWF_Add_c.8:=OWF_Result[8].31;
   		OWF_Result[8].31:=0;
   		OWF_Result[9]:=OWF_Result[9] + 1678588974+OWF_Add_c;
   		OWF_Add_c.9:=OWF_Result[9].31;
   		OWF_Result[9].31:=0;
   		OWF_Result[10]:=OWF_Result[10] + 995137504+OWF_Add_c;
   		OWF_Add_c.10:=OWF_Result[10].31;
   		OWF_Result[10].31:=0;
   		OWF_Result[11]:=OWF_Result[11] + 1432511153+OWF_Add_c;
   		OWF_Add_c.11:=OWF_Result[11].31;
   		OWF_Result[11].31:=0;
   		OWF_Result[12]:=OWF_Result[12] + 148837378+OWF_Add_c;
   		OWF_Add_c.12:=OWF_Result[12].31;
   		OWF_Result[12].31:=0;
   	End_If;
   	If OWF_Input[8].[9] Then
   		OWF_Result[0]:=OWF_Result[0] + 626377956+OWF_Add_c;
   		OWF_Add_c.0:=OWF_Result[0].31;
   		OWF_Result[0].31:=0;
   		OWF_Result[1]:=OWF_Result[1] + 1003201084+OWF_Add_c;
   		OWF_Add_c.1:=OWF_Result[1].31;
   		OWF_Result[1].31:=0;
   		OWF_Result[2]:=OWF_Result[2] + 1213921816+OWF_Add_c;
   		OWF_Add_c.2:=OWF_Result[2].31;
   		OWF_Result[2].31:=0;
   		OWF_Result[3]:=OWF_Result[3] + 637468597+OWF_Add_c;
   		OWF_Add_c.3:=OWF_Result[3].31;
   		OWF_Result[3].31:=0;
   		OWF_Result[4]:=OWF_Result[4] + 1473694468+OWF_Add_c;
   		OWF_Add_c.4:=OWF_Result[4].31;
   		OWF_Result[4].31:=0;
   		OWF_Result[5]:=OWF_Result[5] + 1721369524+OWF_Add_c;
   		OWF_Add_c.5:=OWF_Result[5].31;
   		OWF_Result[5].31:=0;
   		OWF_Result[6]:=OWF_Result[6] + 363430220+OWF_Add_c;
   		OWF_Add_c.6:=OWF_Result[6].31;
   		OWF_Result[6].31:=0;
   		OWF_Result[7]:=OWF_Result[7] + 2083057867+OWF_Add_c;
   		OWF_Add_c.7:=OWF_Result[7].31;
   		OWF_Result[7].31:=0;
   		OWF_Result[8]:=OWF_Result[8] + 994956060+OWF_Add_c;
   		OWF_Add_c.8:=OWF_Result[8].31;
   		OWF_Result[8].31:=0;
   		OWF_Result[9]:=OWF_Result[9] + 1352193715+OWF_Add_c;
   		OWF_Add_c.9:=OWF_Result[9].31;
   		OWF_Result[9].31:=0;
   		OWF_Result[10]:=OWF_Result[10] + 2086908124+OWF_Add_c;
   		OWF_Add_c.10:=OWF_Result[10].31;
   		OWF_Result[10].31:=0;
   		OWF_Result[11]:=OWF_Result[11] + 918226934+OWF_Add_c;
   		OWF_Add_c.11:=OWF_Result[11].31;
   		OWF_Result[11].31:=0;
   		OWF_Result[12]:=OWF_Result[12] + 1905645859+OWF_Add_c;
   		OWF_Add_c.12:=OWF_Result[12].31;
   		OWF_Result[12].31:=0;
   	End_If;
   	If OWF_Input[8].[10] Then
   		OWF_Result[0]:=OWF_Result[0] + 2108694564+OWF_Add_c;
   		OWF_Add_c.0:=OWF_Result[0].31;
   		OWF_Result[0].31:=0;
   		OWF_Result[1]:=OWF_Result[1] + 308494892+OWF_Add_c;
   		OWF_Add_c.1:=OWF_Result[1].31;
   		OWF_Result[1].31:=0;
   		OWF_Result[2]:=OWF_Result[2] + 222147665+OWF_Add_c;
   		OWF_Add_c.2:=OWF_Result[2].31;
   		OWF_Result[2].31:=0;
   		OWF_Result[3]:=OWF_Result[3] + 1066021694+OWF_Add_c;
   		OWF_Add_c.3:=OWF_Result[3].31;
   		OWF_Result[3].31:=0;
   		OWF_Result[4]:=OWF_Result[4] + 735941822+OWF_Add_c;
   		OWF_Add_c.4:=OWF_Result[4].31;
   		OWF_Result[4].31:=0;
   		OWF_Result[5]:=OWF_Result[5] + 1330527490+OWF_Add_c;